   "Carrier_14_SpareInput(4_14)" AT %I1067.4 : Bool;   // SPARE INPUT
   "Carrier_14_SpareInput(4_15)" AT %I1067.5 : Bool;   // SPARE INPUT
   "Carrier_14_SpareInput(4_16)" AT %I1067.6 : Bool;   // SPARE INPUT
   "Carrier_14_SpareInput(4_17)" AT %I1067.7 : Bool;   // SPARE INPUT
   "Carrier_14_Slot5_Output" AT %IW1068 : Word;   // SLOT 5 OUTPUT WORD
   "Carrier_14_IRD400_HMI_24VDC_ENABLE" AT %I1068.0 : Bool;   // IRD 400 PANEL HMI 24V DC POWER
   "Carrier_14_FaultLight_LH" AT %I1068.1 : Bool;   // FAULT LIGHT LH
   "Carrier_14_RunLight_LH" AT %I1068.2 : Bool;   // RUN LIGHT LH
   "Carrier_14_FaultLight_RH" AT %I1068.3 : Bool;   // FAULT LIGHT RH
   "Carrier_14_RunLight_RH" AT %I1068.4 : Bool;   // RUN LIGHT RH
   "Carrier_14_SpareOutput(5_5)" AT %I1068.5 : Bool;   // SPARE OUTPUT
   "Carrier_14_SpareOutput(5_6)" AT %I1068.6 : Bool;   // SPARE OUTPUT
   "Carrier_14_SpareOutput(5_7)" AT %I1068.7 : Bool;   // SPARE OUTPUT
   "Carrier_14_ActualSpeed" AT %IW1070 : Word;   // ACTUAL SPEED
   "Carrier_14_CarrierDriveAlarm" AT %IW1072 : Word;   // CARRIER DRIVE ALARM
   "Carrier_14_CarrierDriveWarning" AT %IW1074 : Word;   // CARRIER DRIVE WARNING
   "Carrier_15_Status" AT %IW1100 : Word;   // CARRIER STATUS WORD
   "Carrier_15_Status.0" AT %I1100.0 : Bool;   // HEARTBEAT
   "Carrier_15_Status.1" AT %I1100.1 : Bool;   // MANUAL
   "Carrier_15_Status.2" AT %I1100.2 : Bool;   // IN_AUTO
   "Carrier_15_Status.3" AT %I1100.3 : Bool;   // POSITIONING_COMPLETE
   "Carrier_15_Status.4" AT %I1100.4 : Bool;   // PRODUCTION HOLD
   "Carrier_15_Status.5" AT %I1100.5 : Bool;   // CARRIER MOVING FORWARD
   "Carrier_15_Status.6" AT %I1100.6 : Bool;   // CARRIER MOVING REVERSE
   "Carrier_15_Status.7" AT %I1100.7 : Bool;   // CARRIER FAULT
   "Carrier_15_Status.8" AT %I1101.0 : Bool;   // CRASH DETECT TRIPPED
   "Carrier_15_Status.9" AT %I1101.1 : Bool;
   "Carrier_15_Status.10" AT %I1101.2 : Bool;
   "Carrier_15_Status.11" AT %I1101.3 : Bool;
   "Carrier_15_Status.12" AT %I1101.4 : Bool;
   "Carrier_15_Status.13" AT %I1101.5 : Bool;
   "Carrier_15_Status.14" AT %I1101.6 : Bool;
   "Carrier_15_Status.15" AT %I1101.7 : Bool;
   "Carrier_15_SDCFaultCode" AT %IW1102 : Word;   // SDC FAULT CODE
   "Carrier_15_CarrierPosition" AT %ID1104 : DWord;   // CARRIER POSITION
   "Carrier_15_CarrierNumber" AT %IW1108 : Word;   // CARRIER NUMBER
   "Carrier_15_G120DControlWord" AT %IW1111 : Word;   // G120D_STW1_CONTROL
   "Carrier_15_G120DControlWord.0" AT %I1111.0 : Bool;   // Bit_00_ON
   "Carrier_15_G120DControlWord.1" AT %I1111.1 : Bool;   // Bit_01_AUS2_INH
   "Carrier_15_G120DControlWord.2" AT %I1111.2 : Bool;   // Bit_02_AUS3_STOP
   "Carrier_15_G120DControlWord.3" AT %I1111.3 : Bool;   // Bit_03_EN
   "Carrier_15_G120DControlWord.4" AT %I1111.4 : Bool;   // Bit_04_EN_RAMP
   "Carrier_15_G120DControlWord.5" AT %I1111.5 : Bool;   // Bit_05_START_RAMP
   "Carrier_15_G120DControlWord.6" AT %I1111.6 : Bool;   // Bit_06_SETPOINT
   "Carrier_15_G120DControlWord.7" AT %I1111.7 : Bool;   // Bit_07_RESET
   "Carrier_15_G120DControlWord.8" AT %I1111.0 : Bool;   // Bit_08_JOG_R
   "Carrier_15_G120DControlWord.9" AT %I1111.1 : Bool;   // Bit_09_JOG_L
   "Carrier_15_G120DControlWord.10" AT %I1111.2 : Bool;   // Bit_10_CONTR_PLC
   "Carrier_15_G120DControlWord.11" AT %I1111.3 : Bool;   // Bit_11_REVERSE
   "Carrier_15_G120DControlWord.12" AT %I1111.4 : Bool;   // Bit_12_BRAKE_RELEASE
   "Carrier_15_G120DControlWord.13" AT %I1111.5 : Bool;   // Bit_13_DDS
   "Carrier_15_G120DControlWord.14" AT %I1111.6 : Bool;   // Bit_14_DO0
   "Carrier_15_G120DControlWord.15" AT %I1111.7 : Bool;   // Bit_15_DO1
   "Carrier_15_G120DStatusWord" AT %IW1112 : Word;   // G120D_ZSW1_STATUS
   "Carrier_15_G120DStatusWord.0" AT %I1112.0 : Bool;   // Bit_00_READY_RUN
   "Carrier_15_G120DStatusWord.1" AT %I1112.1 : Bool;   // Bit_01_READY_ON
   "Carrier_15_G120DStatusWord.2" AT %I1112.2 : Bool;   // Bit_02_ENABLE
   "Carrier_15_G120DStatusWord.3" AT %I1112.3 : Bool;   // Bit_03_FAULT
   "Carrier_15_G120DStatusWord.4" AT %I1112.4 : Bool;   // Bit_04_OFF2
   "Carrier_15_G120DStatusWord.5" AT %I1112.5 : Bool;   // Bit_05_OFF3
   "Carrier_15_G120DStatusWord.6" AT %I1112.6 : Bool;   // Bit_06_LOCK_OUT
   "Carrier_15_G120DStatusWord.7" AT %I1112.7 : Bool;   // Bit_07_WARN
   "Carrier_15_G120DStatusWord.8" AT %I1113.0 : Bool;   // Bit_08_NO_DEVIATION
   "Carrier_15_G120DStatusWord.9" AT %I1113.1 : Bool;   // Bit_09_CONTR_PLC
   "Carrier_15_G120DStatusWord.10" AT %I1113.2 : Bool;   // Bit_10_F_MAX
   "Carrier_15_G120DStatusWord.11" AT %I1113.3 : Bool;   // Bit_11_LIMIT_REACHED
   "Carrier_15_G120DStatusWord.12" AT %I1113.4 : Bool;   // Bit_12_BRAKE_OPEN
   "Carrier_15_G120DStatusWord.13" AT %I1113.5 : Bool;   // Bit_13_NO_OVERTEMP
   "Carrier_15_G120DStatusWord.14" AT %I1113.6 : Bool;   // Bit_14_CW_CCW
   "Carrier_15_G120DStatusWord.15" AT %I1113.7 : Bool;   // Bit_15_OVERL
   "Carrier_15_Slot2_Input" AT %IW1114 : Word;   // SLOT 2 INPUT WORD
   "Carrier_15_CrashDetectSW" AT %I1114.0 : Bool;   // CRASH DETECT SW
   "Carrier_15_SpareSafetyInput(2_1)" AT %I1114.1 : Bool;   // SPARE SAFETY INPUT
   "Carrier_15_SpareSafetyInput(2_2)" AT %I1114.2 : Bool;   // SPARE SAFETY INPUT
   "Carrier_15_SpareSafetyInput(2_3)" AT %I1114.3 : Bool;   // SPARE SAFETY INPUT
   "Carrier_15_SpareSafetyInput(2_4)" AT %I1114.4 : Bool;   // SPARE SAFETY INPUT
   "Carrier_15_SpareSafetyInput(2_5)" AT %I1114.5 : Bool;   // SPARE SAFETY INPUT
   "Carrier_15_SpareSafetyInput(2_6)" AT %I1114.6 : Bool;   // SPARE SAFETY INPUT
   "Carrier_15_SpareSafetyInput(2_7)" AT %I1114.7 : Bool;   // SPARE SAFETY INPUT
   "Carrier_15_Slot3_SafetyOutput" AT %IW1115 : Word;   // SLOT 3 SAFETY OUTPUT WORD
   "Carrier_15_Crash_Detect_OK" AT %I1115.0 : Bool;   // CARRIER CRASH DETECT
   "Carrier_15_SpareSafetyOutput(3_1)" AT %I1115.1 : Bool;   // SPARE SAFETY OUTPUT
   "Carrier_15_SpareSafetyOutput(3_2)" AT %I1115.2 : Bool;   // SPARE SAFETY OUTPUT
   "Carrier_15_SpareSafetyOutput(3_3)" AT %I1115.3 : Bool;   // SPARE SAFETY OUTPUT
   "Carrier_15_SpareSafetyOutput(3_4)" AT %I1115.4 : Bool;   // SPARE SAFETY OUTPUT
   "Carrier_15_SpareSafetyOutput(3_5)" AT %I1115.5 : Bool;   // SPARE SAFETY OUTPUT
   "Carrier_15_SpareSafetyOutput(3_6)" AT %I1115.6 : Bool;   // SPARE SAFETY OUTPUT
   "Carrier_15_SpareSafetyOutput(3_7)" AT %I1115.7 : Bool;   // SPARE SAFETY OUTPUT
   "Carrier_15_Slot4_Input" AT %IW1116 : Word;   // SLOT 4 INPUT WORD
   "Carrier_15_480VPowerOn_MDCB1" AT %I1116.0 : Bool;   // 480 VAC POWER ON MDCB 1
   "Carrier_15_SpareInput(4_1)" AT %I1116.1 : Bool;   // SPARE INPUT
   "Carrier_15_SpareInput(4_2)" AT %I1116.2 : Bool;   // SPARE INPUT
   "Carrier_15_SitopSelectStatus" AT %I1116.3 : Bool;   // SITOP SELECT STATUS
   "Carrier_15_DCsupplyOnPSCB2" AT %I1116.4 : Bool;   // DC SUPPLY ON PSCB 2
   "Carrier_15_SpareInput(4_5)" AT %I1116.5 : Bool;   // SPARE INPUT
   "Carrier_15_SpareInput(4_6)" AT %I1116.6 : Bool;   // SPARE INPUT
   "Carrier_15_SpareInput(4_7)" AT %I1116.7 : Bool;   // SPARE INPUT
   "Carrier_15_PB1_ProdHoldLH" AT %I1117.0 : Bool;   // PB 1 PRODUCTION HOLD LH
   "Carrier_15_PB2_ResetLH" AT %I1117.1 : Bool;   // PB 2 RESET LH
   "Carrier_15_PB3_ProdHoldRH" AT %I1117.2 : Bool;   // PB 3 PRODUCTION HOLD RH
   "Carrier_15_PB4_ResetRH" AT %I1117.3 : Bool;   // PB 4 RESET RH
   "Carrier_15_SpareInput(4_14)" AT %I1117.4 : Bool;   // SPARE INPUT
   "Carrier_15_SpareInput(4_15)" AT %I1117.5 : Bool;   // SPARE INPUT
   "Carrier_15_SpareInput(4_16)" AT %I1117.6 : Bool;   // SPARE INPUT
   "Carrier_15_SpareInput(4_17)" AT %I1117.7 : Bool;   // SPARE INPUT
   "Carrier_15_Slot5_Output" AT %IW1118 : Word;   // SLOT 5 OUTPUT WORD
   "Carrier_15_IRD400_HMI_24VDC_ENABLE" AT %I1118.0 : Bool;   // IRD 400 PANEL HMI 24V DC POWER
   "Carrier_15_FaultLight_LH" AT %I1118.1 : Bool;   // FAULT LIGHT LH
   "Carrier_15_RunLight_LH" AT %I1118.2 : Bool;   // RUN LIGHT LH
   "Carrier_15_FaultLight_RH" AT %I1118.3 : Bool;   // FAULT LIGHT RH
   "Carrier_15_RunLight_RH" AT %I1118.4 : Bool;   // RUN LIGHT RH
   "Carrier_15_SpareOutput(5_5)" AT %I1118.5 : Bool;   // SPARE OUTPUT
   "Carrier_15_SpareOutput(5_6)" AT %I1118.6 : Bool;   // SPARE OUTPUT
   "Carrier_15_SpareOutput(5_7)" AT %I1118.7 : Bool;   // SPARE OUTPUT
   "Carrier_15_ActualSpeed" AT %IW1120 : Word;   // ACTUAL SPEED
   "Carrier_15_CarrierDriveAlarm" AT %IW1122 : Word;   // CARRIER DRIVE ALARM
   "Carrier_15_CarrierDriveWarning" AT %IW1124 : Word;   // CARRIER DRIVE WARNING
   "Carrier_16_Status" AT %IW1150 : Word;   // CARRIER STATUS WORD
   "Carrier_16_Status.0" AT %I1150.0 : Bool;   // HEARTBEAT
   "Carrier_16_Status.1" AT %I1150.1 : Bool;   // MANUAL
   "Carrier_16_Status.2" AT %I1150.2 : Bool;   // IN_AUTO
   "Carrier_16_Status.3" AT %I1150.3 : Bool;   // POSITIONING_COMPLETE
   "Carrier_16_Status.4" AT %I1150.4 : Bool;   // PRODUCTION HOLD
   "Carrier_16_Status.5" AT %I1150.5 : Bool;   // CARRIER MOVING FORWARD
   "Carrier_16_Status.6" AT %I1150.6 : Bool;   // CARRIER MOVING REVERSE
   "Carrier_16_Status.7" AT %I1150.7 : Bool;   // CARRIER FAULT
   "Carrier_16_Status.8" AT %I1151.0 : Bool;   // CRASH DETECT TRIPPED
   "Carrier_16_Status.9" AT %I1151.1 : Bool;
   "Carrier_16_Status.10" AT %I1151.2 : Bool;
   "Carrier_16_Status.11" AT %I1151.3 : Bool;
   "Carrier_16_Status.12" AT %I1151.4 : Bool;
   "Carrier_16_Status.13" AT %I1151.5 : Bool;
   "Carrier_16_Status.14" AT %I1151.6 : Bool;
   "Carrier_16_Status.15" AT %I1151.7 : Bool;
   "Carrier_16_SDCFaultCode" AT %IW1152 : Word;   // SDC FAULT CODE
   "Carrier_16_CarrierPosition" AT %ID1154 : DWord;   // CARRIER POSITION
   "Carrier_16_CarrierNumber" AT %IW1158 : Word;   // CARRIER NUMBER
   "Carrier_16_G120DControlWord" AT %IW1160 : Word;   // G120D_STW1_CONTROL
   "Carrier_16_G120DControlWord.0" AT %I1160.0 : Bool;   // Bit_00_ON
   "Carrier_16_G120DControlWord.1" AT %I1160.1 : Bool;   // Bit_01_AUS2_INH
   "Carrier_16_G120DControlWord.2" AT %I1160.2 : Bool;   // Bit_02_AUS3_STOP
   "Carrier_16_G120DControlWord.3" AT %I1160.3 : Bool;   // Bit_03_EN
   "Carrier_16_G120DControlWord.4" AT %I1160.4 : Bool;   // Bit_04_EN_RAMP
   "Carrier_16_G120DControlWord.5" AT %I1160.5 : Bool;   // Bit_05_START_RAMP
   "Carrier_16_G120DControlWord.6" AT %I1160.6 : Bool;   // Bit_06_SETPOINT
   "Carrier_16_G120DControlWord.7" AT %I1160.7 : Bool;   // Bit_07_RESET
   "Carrier_16_G120DControlWord.8" AT %I1161.0 : Bool;   // Bit_08_JOG_R
   "Carrier_16_G120DControlWord.9" AT %I1161.1 : Bool;   // Bit_09_JOG_L
   "Carrier_16_G120DControlWord.10" AT %I1161.2 : Bool;   // Bit_10_CONTR_PLC
   "Carrier_16_G120DControlWord.11" AT %I1161.3 : Bool;   // Bit_11_REVERSE
   "Carrier_16_G120DControlWord.12" AT %I1161.4 : Bool;   // Bit_12_BRAKE_RELEASE
   "Carrier_16_G120DControlWord.13" AT %I1161.5 : Bool;   // Bit_13_DDS
   "Carrier_16_G120DControlWord.14" AT %I1161.6 : Bool;   // Bit_14_DO0
   "Carrier_16_G120DControlWord.15" AT %I1161.7 : Bool;   // Bit_15_DO1
   "Carrier_16_G120DStatusWord" AT %IW1162 : Word;   // G120D_ZSW1_STATUS
   "Carrier_16_G120DStatusWord.0" AT %I1162.0 : Bool;   // Bit_00_READY_RUN
   "Carrier_16_G120DStatusWord.1" AT %I1162.1 : Bool;   // Bit_01_READY_ON
   "Carrier_16_G120DStatusWord.2" AT %I1162.2 : Bool;   // Bit_02_ENABLE
   "Carrier_16_G120DStatusWord.3" AT %I1162.3 : Bool;   // Bit_03_FAULT
   "Carrier_16_G120DStatusWord.4" AT %I1162.4 : Bool;   // Bit_04_OFF2
   "Carrier_16_G120DStatusWord.5" AT %I1162.5 : Bool;   // Bit_05_OFF3
   "Carrier_16_G120DStatusWord.6" AT %I1162.6 : Bool;   // Bit_06_LOCK_OUT
   "Carrier_16_G120DStatusWord.7" AT %I1162.7 : Bool;   // Bit_07_WARN
   "Carrier_16_G120DStatusWord.8" AT %I1163.0 : Bool;   // Bit_08_NO_DEVIATION
   "Carrier_16_G120DStatusWord.9" AT %I1163.1 : Bool;   // Bit_09_CONTR_PLC
   "Carrier_16_G120DStatusWord.10" AT %I1163.2 : Bool;   // Bit_10_F_MAX
   "Carrier_16_G120DStatusWord.11" AT %I1163.3 : Bool;   // Bit_11_LIMIT_REACHED
   "Carrier_16_G120DStatusWord.12" AT %I1163.4 : Bool;   // Bit_12_BRAKE_OPEN
   "Carrier_16_G120DStatusWord.13" AT %I1163.5 : Bool;   // Bit_13_NO_OVERTEMP
   "Carrier_16_G120DStatusWord.14" AT %I1163.6 : Bool;   // Bit_14_CW_CCW
   "Carrier_16_G120DStatusWord.15" AT %I1163.7 : Bool;   // Bit_15_OVERL
   "Carrier_16_Slot2_Input" AT %IW1164 : Word;   // SLOT 2 INPUT WORD
   "Carrier_16_CrashDetectSW" AT %I1164.0 : Bool;   // CRASH DETECT SW
   "Carrier_16_SpareSafetyInput(2_1)" AT %I1164.1 : Bool;   // SPARE SAFETY INPUT
   "Carrier_16_SpareSafetyInput(2_2)" AT %I1164.2 : Bool;   // SPARE SAFETY INPUT
   "Carrier_16_SpareSafetyInput(2_3)" AT %I1164.3 : Bool;   // SPARE SAFETY INPUT
   "Carrier_16_SpareSafetyInput(2_4)" AT %I1164.4 : Bool;   // SPARE SAFETY INPUT
   "Carrier_16_SpareSafetyInput(2_5)" AT %I1164.5 : Bool;   // SPARE SAFETY INPUT
   "Carrier_16_SpareSafetyInput(2_6)" AT %I1164.6 : Bool;   // SPARE SAFETY INPUT
   "Carrier_16_SpareSafetyInput(2_7)" AT %I1164.7 : Bool;   // SPARE SAFETY INPUT
   "Carrier_16_Slot3_SafetyOutput" AT %IW1165 : Word;   // SLOT 3 SAFETY OUTPUT WORD
   "Carrier_16_Crash_Detect_OK" AT %I1165.0 : Bool;   // CARRIER CRASH DETECT
   "Carrier_16_SpareSafetyOutput(3_1)" AT %I1165.1 : Bool;   // SPARE SAFETY OUTPUT
   "Carrier_16_SpareSafetyOutput(3_2)" AT %I1165.2 : Bool;   // SPARE SAFETY OUTPUT
   "Carrier_16_SpareSafetyOutput(3_3)" AT %I1165.3 : Bool;   // SPARE SAFETY OUTPUT
   "Carrier_16_SpareSafetyOutput(3_4)" AT %I1165.4 : Bool;   // SPARE SAFETY OUTPUT
   "Carrier_16_SpareSafetyOutput(3_5)" AT %I1165.5 : Bool;   // SPARE SAFETY OUTPUT
   "Carrier_16_SpareSafetyOutput(3_6)" AT %I1165.6 : Bool;   // SPARE SAFETY OUTPUT
   "Carrier_16_SpareSafetyOutput(3_7)" AT %I1165.7 : Bool;   // SPARE SAFETY OUTPUT
   "Carrier_16_Slot4_Input" AT %IW1166 : Word;   // SLOT 4 INPUT WORD
   "Carrier_16_480VPowerOn_MDCB1" AT %I1166.0 : Bool;   // 480 VAC POWER ON MDCB 1
   "Carrier_16_SpareInput(4_1)" AT %I1166.1 : Bool;   // SPARE INPUT
   "Carrier_16_SpareInput(4_2)" AT %I1166.2 : Bool;   // SPARE INPUT
   "Carrier_16_SitopSelectStatus" AT %I1166.3 : Bool;   // SITOP SELECT STATUS
   "Carrier_16_DCsupplyOnPSCB2" AT %I1166.4 : Bool;   // DC SUPPLY ON PSCB 2
   "Carrier_16_SpareInput(4_5)" AT %I1166.5 : Bool;   // SPARE INPUT
   "Carrier_16_SpareInput(4_6)" AT %I1166.6 : Bool;   // SPARE INPUT
   "Carrier_16_SpareInput(4_7)" AT %I1166.7 : Bool;   // SPARE INPUT
   "Carrier_16_PB1_ProdHoldLH" AT %I1167.0 : Bool;   // PB 1 PRODUCTION HOLD LH
   "Carrier_16_PB2_ResetLH" AT %I1167.1 : Bool;   // PB 2 RESET LH
   "Carrier_16_PB3_ProdHoldRH" AT %I1167.2 : Bool;   // PB 3 PRODUCTION HOLD RH
   "Carrier_16_PB4_ResetRH" AT %I1167.3 : Bool;   // PB 4 RESET RH
   "Carrier_16_SpareInput(4_14)" AT %I1167.4 : Bool;   // SPARE INPUT
   "Carrier_16_SpareInput(4_15)" AT %I1167.5 : Bool;   // SPARE INPUT
   "Carrier_16_SpareInput(4_16)" AT %I1167.6 : Bool;   // SPARE INPUT
   "Carrier_16_SpareInput(4_17)" AT %I1167.7 : Bool;   // SPARE INPUT
   "Carrier_16_Slot5_Output" AT %IW1168 : Word;   // SLOT 5 OUTPUT WORD
   "Carrier_16_IRD400_HMI_24VDC_ENABLE" AT %I1168.0 : Bool;   // IRD 400 PANEL HMI 24V DC POWER
   "Carrier_16_FaultLight_LH" AT %I1168.1 : Bool;   // FAULT LIGHT LH
   "Carrier_16_RunLight_LH" AT %I1168.2 : Bool;   // RUN LIGHT LH
   "Carrier_16_FaultLight_RH" AT %I1168.3 : Bool;   // FAULT LIGHT RH
   "Carrier_16_RunLight_RH" AT %I1168.4 : Bool;   // RUN LIGHT RH
   "Carrier_16_SpareOutput(5_5)" AT %I1168.5 : Bool;   // SPARE OUTPUT
   "Carrier_16_SpareOutput(5_6)" AT %I1168.6 : Bool;   // SPARE OUTPUT
   "Carrier_16_SpareOutput(5_7)" AT %I1168.7 : Bool;   // SPARE OUTPUT
   "Carrier_16_ActualSpeed" AT %IW1170 : Word;   // ACTUAL SPEED
   "Carrier_16_CarrierDriveAlarm" AT %IW1172 : Word;   // CARRIER DRIVE ALARM
   "Carrier_16_CarrierDriveWarning" AT %IW1174 : Word;   // CARRIER DRIVE WARNING
   "Carrier_17_Status" AT %IW1200 : Word;   // CARRIER STATUS WORD
   "Carrier_17_Status.0" AT %I1200.0 : Bool;   // HEARTBEAT
   "Carrier_17_Status.1" AT %I1200.1 : Bool;   // MANUAL
   "Carrier_17_Status.2" AT %I1200.2 : Bool;   // IN_AUTO
   "Carrier_17_Status.3" AT %I1200.3 : Bool;   // POSITIONING_COMPLETE
   "Carrier_17_Status.4" AT %I1200.4 : Bool;   // PRODUCTION HOLD
   "Carrier_17_Status.5" AT %I1200.5 : Bool;   // CARRIER MOVING FORWARD
   "Carrier_17_Status.6" AT %I1200.6 : Bool;   // CARRIER MOVING REVERSE
   "Carrier_17_Status.7" AT %I1200.7 : Bool;   // CARRIER FAULT
   "Carrier_17_Status.8" AT %I1201.0 : Bool;   // CRASH DETECT TRIPPED
   "Carrier_17_Status.9" AT %I1201.1 : Bool;
   "Carrier_17_Status.10" AT %I1201.2 : Bool;
   "Carrier_17_Status.11" AT %I1201.3 : Bool;
   "Carrier_17_Status.12" AT %I1201.4 : Bool;
   "Carrier_17_Status.13" AT %I1201.5 : Bool;
   "Carrier_17_Status.14" AT %I1201.6 : Bool;
   "Carrier_17_Status.15" AT %I1201.7 : Bool;
   "Carrier_17_SDCFaultCode" AT %IW1202 : Word;   // SDC FAULT CODE
   "Carrier_17_CarrierPosition" AT %ID1204 : DWord;   // CARRIER POSITION
   "Carrier_17_CarrierNumber" AT %IW1208 : Word;   // CARRIER NUMBER
   "Carrier_17_G120DControlWord" AT %IW1212 : Word;   // G120D_STW1_CONTROL
   "Carrier_17_G120DControlWord.0" AT %I1212.0 : Bool;   // Bit_00_ON
   "Carrier_17_G120DControlWord.1" AT %I1212.1 : Bool;   // Bit_01_AUS2_INH
   "Carrier_17_G120DControlWord.2" AT %I1212.2 : Bool;   // Bit_02_AUS3_STOP
   "Carrier_17_G120DControlWord.3" AT %I1212.3 : Bool;   // Bit_03_EN
   "Carrier_17_G120DControlWord.4" AT %I1212.4 : Bool;   // Bit_04_EN_RAMP
   "Carrier_17_G120DControlWord.5" AT %I1212.5 : Bool;   // Bit_05_START_RAMP
   "Carrier_17_G120DControlWord.6" AT %I1212.6 : Bool;   // Bit_06_SETPOINT
   "Carrier_17_G120DControlWord.7" AT %I1212.7 : Bool;   // Bit_07_RESET
   "Carrier_17_G120DControlWord.8" AT %I1212.0 : Bool;   // Bit_08_JOG_R
   "Carrier_17_G120DControlWord.9" AT %I1212.1 : Bool;   // Bit_09_JOG_L
   "Carrier_17_G120DControlWord.10" AT %I1212.2 : Bool;   // Bit_10_CONTR_PLC
   "Carrier_17_G120DControlWord.11" AT %I1212.3 : Bool;   // Bit_11_REVERSE
   "Carrier_17_G120DControlWord.12" AT %I1212.4 : Bool;   // Bit_12_BRAKE_RELEASE
   "Carrier_17_G120DControlWord.13" AT %I1212.5 : Bool;   // Bit_13_DDS
   "Carrier_17_G120DControlWord.14" AT %I1212.6 : Bool;   // Bit_14_DO0
   "Carrier_17_G120DControlWord.15" AT %I1212.7 : Bool;   // Bit_15_DO1
   "Carrier_17_G120DStatusWord" AT %IW1212 : Word;   // G120D_ZSW1_STATUS
   "Carrier_17_G120DStatusWord.0" AT %I1212.0 : Bool;   // Bit_00_READY_RUN
   "Carrier_17_G120DStatusWord.1" AT %I1212.1 : Bool;   // Bit_01_READY_ON
   "Carrier_17_G120DStatusWord.2" AT %I1212.2 : Bool;   // Bit_02_ENABLE
   "Carrier_17_G120DStatusWord.3" AT %I1212.3 : Bool;   // Bit_03_FAULT
   "Carrier_17_G120DStatusWord.4" AT %I1212.4 : Bool;   // Bit_04_OFF2
   "Carrier_17_G120DStatusWord.5" AT %I1212.5 : Bool;   // Bit_05_OFF3
   "Carrier_17_G120DStatusWord.6" AT %I1212.6 : Bool;   // Bit_06_LOCK_OUT
   "Carrier_17_G120DStatusWord.7" AT %I1212.7 : Bool;   // Bit_07_WARN
   "Carrier_17_G120DStatusWord.8" AT %I1213.0 : Bool;   // Bit_08_NO_DEVIATION
   "Carrier_17_G120DStatusWord.9" AT %I1213.1 : Bool;   // Bit_09_CONTR_PLC
   "Carrier_17_G120DStatusWord.10" AT %I1213.2 : Bool;   // Bit_10_F_MAX
   "Carrier_17_G120DStatusWord.11" AT %I1213.3 : Bool;   // Bit_11_LIMIT_REACHED
   "Carrier_17_G120DStatusWord.12" AT %I1213.4 : Bool;   // Bit_12_BRAKE_OPEN
   "Carrier_17_G120DStatusWord.13" AT %I1213.5 : Bool;   // Bit_13_NO_OVERTEMP
   "Carrier_17_G120DStatusWord.14" AT %I1213.6 : Bool;   // Bit_14_CW_CCW
   "Carrier_17_G120DStatusWord.15" AT %I1213.7 : Bool;   // Bit_15_OVERL
   "Carrier_17_Slot2_Input" AT %IW1214 : Word;   // SLOT 2 INPUT WORD
   "Carrier_17_CrashDetectSW" AT %I1214.0 : Bool;   // CRASH DETECT SW
   "Carrier_17_SpareSafetyInput(2_1)" AT %I1214.1 : Bool;   // SPARE SAFETY INPUT
   "Carrier_17_SpareSafetyInput(2_2)" AT %I1214.2 : Bool;   // SPARE SAFETY INPUT
   "Carrier_17_SpareSafetyInput(2_3)" AT %I1214.3 : Bool;   // SPARE SAFETY INPUT
   "Carrier_17_SpareSafetyInput(2_4)" AT %I1214.4 : Bool;   // SPARE SAFETY INPUT
   "Carrier_17_SpareSafetyInput(2_5)" AT %I1214.5 : Bool;   // SPARE SAFETY INPUT
   "Carrier_17_SpareSafetyInput(2_6)" AT %I1214.6 : Bool;   // SPARE SAFETY INPUT
   "Carrier_17_SpareSafetyInput(2_7)" AT %I1214.7 : Bool;   // SPARE SAFETY INPUT
   "Carrier_17_Slot3_SafetyOutput" AT %IW1215 : Word;   // SLOT 3 SAFETY OUTPUT WORD
   "Carrier_17_Crash_Detect_OK" AT %I1215.0 : Bool;   // CARRIER CRASH DETECT
   "Carrier_17_SpareSafetyOutput(3_1)" AT %I1215.1 : Bool;   // SPARE SAFETY OUTPUT
   "Carrier_17_SpareSafetyOutput(3_2)" AT %I1215.2 : Bool;   // SPARE SAFETY OUTPUT
   "Carrier_17_SpareSafetyOutput(3_3)" AT %I1215.3 : Bool;   // SPARE SAFETY OUTPUT
   "Carrier_17_SpareSafetyOutput(3_4)" AT %I1215.4 : Bool;   // SPARE SAFETY OUTPUT
   "Carrier_17_SpareSafetyOutput(3_5)" AT %I1215.5 : Bool;   // SPARE SAFETY OUTPUT
   "Carrier_17_SpareSafetyOutput(3_6)" AT %I1215.6 : Bool;   // SPARE SAFETY OUTPUT
   "Carrier_17_SpareSafetyOutput(3_7)" AT %I1215.7 : Bool;   // SPARE SAFETY OUTPUT
   "Carrier_17_Slot4_Input" AT %IW1216 : Word;   // SLOT 4 INPUT WORD
   "Carrier_17_480VPowerOn_MDCB1" AT %I1216.0 : Bool;   // 480 VAC POWER ON MDCB 1
   "Carrier_17_SpareInput(4_1)" AT %I1216.1 : Bool;   // SPARE INPUT
   "Carrier_17_SpareInput(4_2)" AT %I1216.2 : Bool;   // SPARE INPUT
   "Carrier_17_SitopSelectStatus" AT %I1216.3 : Bool;   // SITOP SELECT STATUS
   "Carrier_17_DCsupplyOnPSCB2" AT %I1216.4 : Bool;   // DC SUPPLY ON PSCB 2
   "Carrier_17_SpareInput(4_5)" AT %I1216.5 : Bool;   // SPARE INPUT
   "Carrier_17_SpareInput(4_6)" AT %I1216.6 : Bool;   // SPARE INPUT
   "Carrier_17_SpareInput(4_7)" AT %I1216.7 : Bool;   // SPARE INPUT
   "Carrier_17_PB1_ProdHoldLH" AT %I1217.0 : Bool;   // PB 1 PRODUCTION HOLD LH
   "Carrier_17_PB2_ResetLH" AT %I1217.1 : Bool;   // PB 2 RESET LH
   "Carrier_17_PB3_ProdHoldRH" AT %I1217.2 : Bool;   // PB 3 PRODUCTION HOLD RH
   "Carrier_17_PB4_ResetRH" AT %I1217.3 : Bool;   // PB 4 RESET RH
   "Carrier_17_SpareInput(4_14)" AT %I1217.4 : Bool;   // SPARE INPUT
   "Carrier_17_SpareInput(4_15)" AT %I1217.5 : Bool;   // SPARE INPUT
   "Carrier_17_SpareInput(4_16)" AT %I1217.6 : Bool;   // SPARE INPUT
   "Carrier_17_SpareInput(4_17)" AT %I1217.7 : Bool;   // SPARE INPUT
   "Carrier_17_Slot5_Output" AT %IW1218 : Word;   // SLOT 5 OUTPUT WORD
   "Carrier_17_IRD400_HMI_24VDC_ENABLE" AT %I1218.0 : Bool;   // IRD 400 PANEL HMI 24V DC POWER
   "Carrier_17_FaultLight_LH" AT %I1218.1 : Bool;   // FAULT LIGHT LH
   "Carrier_17_RunLight_LH" AT %I1218.2 : Bool;   // RUN LIGHT LH
   "Carrier_17_FaultLight_RH" AT %I1218.3 : Bool;   // FAULT LIGHT RH
   "Carrier_17_RunLight_RH" AT %I1218.4 : Bool;   // RUN LIGHT RH
   "Carrier_17_SpareOutput(5_5)" AT %I1218.5 : Bool;   // SPARE OUTPUT
   "Carrier_17_SpareOutput(5_6)" AT %I1218.6 : Bool;   // SPARE OUTPUT
   "Carrier_17_SpareOutput(5_7)" AT %I1218.7 : Bool;   // SPARE OUTPUT
   "Carrier_17_ActualSpeed" AT %IW1220 : Word;   // ACTUAL SPEED
   "Carrier_17_CarrierDriveAlarm" AT %IW1222 : Word;   // CARRIER DRIVE ALARM
   "Carrier_17_CarrierDriveWarning" AT %IW1224 : Word;   // CARRIER DRIVE WARNING
   "Carrier_18_Status" AT %IW1250 : Word;   // CARRIER STATUS WORD
   "Carrier_18_Status.0" AT %I1250.0 : Bool;   // HEARTBEAT
   "Carrier_18_Status.1" AT %I1250.1 : Bool;   // MANUAL
   "Carrier_18_Status.2" AT %I1250.2 : Bool;   // IN_AUTO
   "Carrier_18_Status.3" AT %I1250.3 : Bool;   // POSITIONING_COMPLETE
   "Carrier_18_Status.4" AT %I1250.4 : Bool;   // PRODUCTION HOLD
   "Carrier_18_Status.5" AT %I1250.5 : Bool;   // CARRIER MOVING FORWARD
   "Carrier_18_Status.6" AT %I1250.6 : Bool;   // CARRIER MOVING REVERSE
   "Carrier_18_Status.7" AT %I1250.7 : Bool;   // CARRIER FAULT
   "Carrier_18_Status.8" AT %I1251.0 : Bool;   // CRASH DETECT TRIPPED
   "Carrier_18_Status.9" AT %I1251.1 : Bool;
   "Carrier_18_Status.10" AT %I1251.2 : Bool;
   "Carrier_18_Status.11" AT %I1251.3 : Bool;
   "Carrier_18_Status.12" AT %I1251.4 : Bool;
   "Carrier_18_Status.13" AT %I1251.5 : Bool;
   "Carrier_18_Status.14" AT %I1251.6 : Bool;
   "Carrier_18_Status.15" AT %I1251.7 : Bool;
   "Carrier_18_SDCFaultCode" AT %IW1252 : Word;   // SDC FAULT CODE
   "Carrier_18_CarrierPosition" AT %ID1254 : DWord;   // CARRIER POSITION
   "Carrier_18_CarrierNumber" AT %IW1258 : Word;   // CARRIER NUMBER
   "Carrier_18_G120DControlWord" AT %IW1260 : Word;   // G120D_STW1_CONTROL
   "Carrier_18_G120DControlWord.0" AT %I1260.0 : Bool;   // Bit_00_ON
   "Carrier_18_G120DControlWord.1" AT %I1260.1 : Bool;   // Bit_01_AUS2_INH
   "Carrier_18_G120DControlWord.2" AT %I1260.2 : Bool;   // Bit_02_AUS3_STOP
   "Carrier_18_G120DControlWord.3" AT %I1260.3 : Bool;   // Bit_03_EN
   "Carrier_18_G120DControlWord.4" AT %I1260.4 : Bool;   // Bit_04_EN_RAMP
   "Carrier_18_G120DControlWord.5" AT %I1260.5 : Bool;   // Bit_05_START_RAMP
   "Carrier_18_G120DControlWord.6" AT %I1260.6 : Bool;   // Bit_06_SETPOINT
   "Carrier_18_G120DControlWord.7" AT %I1260.7 : Bool;   // Bit_07_RESET
   "Carrier_18_G120DControlWord.8" AT %I1261.0 : Bool;   // Bit_08_JOG_R
   "Carrier_18_G120DControlWord.9" AT %I1261.1 : Bool;   // Bit_09_JOG_L
   "Carrier_18_G120DControlWord.10" AT %I1261.2 : Bool;   // Bit_10_CONTR_PLC
   "Carrier_18_G120DControlWord.11" AT %I1261.3 : Bool;   // Bit_11_REVERSE
   "Carrier_18_G120DControlWord.12" AT %I1261.4 : Bool;   // Bit_12_BRAKE_RELEASE
   "Carrier_18_G120DControlWord.13" AT %I1261.5 : Bool;   // Bit_13_DDS
   "Carrier_18_G120DControlWord.14" AT %I1261.6 : Bool;   // Bit_14_DO0
   "Carrier_18_G120DControlWord.15" AT %I1261.7 : Bool;   // Bit_15_DO1
   "Carrier_18_G120DStatusWord" AT %IW1262 : Word;   // G120D_ZSW1_STATUS
   "Carrier_18_G120DStatusWord.0" AT %I1262.0 : Bool;   // Bit_00_READY_RUN
   "Carrier_18_G120DStatusWord.1" AT %I1262.1 : Bool;   // Bit_01_READY_ON
   "Carrier_18_G120DStatusWord.2" AT %I1262.2 : Bool;   // Bit_02_ENABLE
   "Carrier_18_G120DStatusWord.3" AT %I1262.3 : Bool;   // Bit_03_FAULT
   "Carrier_18_G120DStatusWord.4" AT %I1262.4 : Bool;   // Bit_04_OFF2
   "Carrier_18_G120DStatusWord.5" AT %I1262.5 : Bool;   // Bit_05_OFF3
   "Carrier_18_G120DStatusWord.6" AT %I1262.6 : Bool;   // Bit_06_LOCK_OUT
   "Carrier_18_G120DStatusWord.7" AT %I1262.7 : Bool;   // Bit_07_WARN
   "Carrier_18_G120DStatusWord.8" AT %I1263.0 : Bool;   // Bit_08_NO_DEVIATION
   "Carrier_18_G120DStatusWord.9" AT %I1263.1 : Bool;   // Bit_09_CONTR_PLC
   "Carrier_18_G120DStatusWord.10" AT %I1263.2 : Bool;   // Bit_10_F_MAX
   "Carrier_18_G120DStatusWord.11" AT %I1263.3 : Bool;   // Bit_11_LIMIT_REACHED
   "Carrier_18_G120DStatusWord.12" AT %I1263.4 : Bool;   // Bit_12_BRAKE_OPEN
   "Carrier_18_G120DStatusWord.13" AT %I1263.5 : Bool;   // Bit_13_NO_OVERTEMP
   "Carrier_18_G120DStatusWord.14" AT %I1263.6 : Bool;   // Bit_14_CW_CCW
   "Carrier_18_G120DStatusWord.15" AT %I1263.7 : Bool;   // Bit_15_OVERL
   "Carrier_18_Slot2_Input" AT %IW1264 : Word;   // SLOT 2 INPUT WORD
   "Carrier_18_CrashDetectSW" AT %I1264.0 : Bool;   // CRASH DETECT SW
   "Carrier_18_SpareSafetyInput(2_1)" AT %I1264.1 : Bool;   // SPARE SAFETY INPUT
   "Carrier_18_SpareSafetyInput(2_2)" AT %I1264.2 : Bool;   // SPARE SAFETY INPUT
   "Carrier_18_SpareSafetyInput(2_3)" AT %I1264.3 : Bool;   // SPARE SAFETY INPUT
   "Carrier_18_SpareSafetyInput(2_4)" AT %I1264.4 : Bool;   // SPARE SAFETY INPUT
   "Carrier_18_SpareSafetyInput(2_5)" AT %I1264.5 : Bool;   // SPARE SAFETY INPUT
   "Carrier_18_SpareSafetyInput(2_6)" AT %I1264.6 : Bool;   // SPARE SAFETY INPUT
   "Carrier_18_SpareSafetyInput(2_7)" AT %I1264.7 : Bool;   // SPARE SAFETY INPUT
   "Carrier_18_Slot3_SafetyOutput" AT %IW1265 : Word;   // SLOT 3 SAFETY OUTPUT WORD
   "Carrier_18_Crash_Detect_OK" AT %I1265.0 : Bool;   // CARRIER CRASH DETECT
   "Carrier_18_SpareSafetyOutput(3_1)" AT %I1265.1 : Bool;   // SPARE SAFETY OUTPUT
   "Carrier_18_SpareSafetyOutput(3_2)" AT %I1265.2 : Bool;   // SPARE SAFETY OUTPUT
   "Carrier_18_SpareSafetyOutput(3_3)" AT %I1265.3 : Bool;   // SPARE SAFETY OUTPUT
   "Carrier_18_SpareSafetyOutput(3_4)" AT %I1265.4 : Bool;   // SPARE SAFETY OUTPUT
   "Carrier_18_SpareSafetyOutput(3_5)" AT %I1265.5 : Bool;   // SPARE SAFETY OUTPUT
   "Carrier_18_SpareSafetyOutput(3_6)" AT %I1265.6 : Bool;   // SPARE SAFETY OUTPUT
   "Carrier_18_SpareSafetyOutput(3_7)" AT %I1265.7 : Bool;   // SPARE SAFETY OUTPUT
   "Carrier_18_Slot4_Input" AT %IW1266 : Word;   // SLOT 4 INPUT WORD
   "Carrier_18_480VPowerOn_MDCB1" AT %I1266.0 : Bool;   // 480 VAC POWER ON MDCB 1
   "Carrier_18_SpareInput(4_1)" AT %I1266.1 : Bool;   // SPARE INPUT
   "Carrier_18_SpareInput(4_2)" AT %I1266.2 : Bool;   // SPARE INPUT
   "Carrier_18_SitopSelectStatus" AT %I1266.3 : Bool;   // SITOP SELECT STATUS
   "Carrier_18_DCsupplyOnPSCB2" AT %I1266.4 : Bool;   // DC SUPPLY ON PSCB 2
   "Carrier_18_SpareInput(4_5)" AT %I1266.5 : Bool;   // SPARE INPUT
   "Carrier_18_SpareInput(4_6)" AT %I1266.6 : Bool;   // SPARE INPUT
   "Carrier_18_SpareInput(4_7)" AT %I1266.7 : Bool;   // SPARE INPUT
   "Carrier_18_PB1_ProdHoldLH" AT %I1267.0 : Bool;   // PB 1 PRODUCTION HOLD LH
   "Carrier_18_PB2_ResetLH" AT %I1267.1 : Bool;   // PB 2 RESET LH
   "Carrier_18_PB3_ProdHoldRH" AT %I1267.2 : Bool;   // PB 3 PRODUCTION HOLD RH
   "Carrier_18_PB4_ResetRH" AT %I1267.3 : Bool;   // PB 4 RESET RH
   "Carrier_18_SpareInput(4_14)" AT %I1267.4 : Bool;   // SPARE INPUT
   "Carrier_18_SpareInput(4_15)" AT %I1267.5 : Bool;   // SPARE INPUT
   "Carrier_18_SpareInput(4_16)" AT %I1267.6 : Bool;   // SPARE INPUT
   "Carrier_18_SpareInput(4_17)" AT %I1267.7 : Bool;   // SPARE INPUT
   "Carrier_18_Slot5_Output" AT %IW1268 : Word;   // SLOT 5 OUTPUT WORD
   "Carrier_18_IRD400_HMI_24VDC_ENABLE" AT %I1268.0 : Bool;   // IRD 400 PANEL HMI 24V DC POWER
   "Carrier_18_FaultLight_LH" AT %I1268.1 : Bool;   // FAULT LIGHT LH
   "Carrier_18_RunLight_LH" AT %I1268.2 : Bool;   // RUN LIGHT LH
   "Carrier_18_FaultLight_RH" AT %I1268.3 : Bool;   // FAULT LIGHT RH
   "Carrier_18_RunLight_RH" AT %I1268.4 : Bool;   // RUN LIGHT RH
   "Carrier_18_SpareOutput(5_5)" AT %I1268.5 : Bool;   // SPARE OUTPUT
   "Carrier_18_SpareOutput(5_6)" AT %I1268.6 : Bool;   // SPARE OUTPUT
   "Carrier_18_SpareOutput(5_7)" AT %I1268.7 : Bool;   // SPARE OUTPUT
   "Carrier_18_ActualSpeed" AT %IW1270 : Word;   // ACTUAL SPEED
   "Carrier_18_CarrierDriveAlarm" AT %IW1272 : Word;   // CARRIER DRIVE ALARM
   "Carrier_18_CarrierDriveWarning" AT %IW1274 : Word;   // CARRIER DRIVE WARNING
   "Carrier_19_Status" AT %IW1300 : Word;   // CARRIER STATUS WORD
   "Carrier_19_Status.0" AT %I1300.0 : Bool;   // HEARTBEAT
   "Carrier_19_Status.1" AT %I1300.1 : Bool;   // MANUAL
   "Carrier_19_Status.2" AT %I1300.2 : Bool;   // IN_AUTO
   "Carrier_19_Status.3" AT %I1300.3 : Bool;   // POSITIONING_COMPLETE
   "Carrier_19_Status.4" AT %I1300.4 : Bool;   // PRODUCTION HOLD
   "Carrier_19_Status.5" AT %I1300.5 : Bool;   // CARRIER MOVING FORWARD
   "Carrier_19_Status.6" AT %I1300.6 : Bool;   // CARRIER MOVING REVERSE
   "Carrier_19_Status.7" AT %I1300.7 : Bool;   // CARRIER FAULT
   "Carrier_19_Status.8" AT %I1301.0 : Bool;   // CRASH DETECT TRIPPED
   "Carrier_19_Status.9" AT %I1301.1 : Bool;
   "Carrier_19_Status.10" AT %I1301.2 : Bool;
   "Carrier_19_Status.11" AT %I1301.3 : Bool;
   "Carrier_19_Status.12" AT %I1301.4 : Bool;
   "Carrier_19_Status.13" AT %I1301.5 : Bool;
   "Carrier_19_Status.14" AT %I1301.6 : Bool;
   "Carrier_19_Status.15" AT %I1301.7 : Bool;
   "Carrier_19_SDCFaultCode" AT %IW1302 : Word;   // SDC FAULT CODE
   "Carrier_19_CarrierPosition" AT %ID1304 : DWord;   // CARRIER POSITION
   "Carrier_19_CarrierNumber" AT %IW1308 : Word;   // CARRIER NUMBER
   "Carrier_19_G120DControlWord" AT %IW1310 : Word;   // G120D_STW1_CONTROL
   "Carrier_19_G120DControlWord.0" AT %I1310.0 : Bool;   // Bit_00_ON
   "Carrier_19_G120DControlWord.1" AT %I1310.1 : Bool;   // Bit_01_AUS2_INH
   "Carrier_19_G120DControlWord.2" AT %I1310.2 : Bool;   // Bit_02_AUS3_STOP
   "Carrier_19_G120DControlWord.3" AT %I1310.3 : Bool;   // Bit_03_EN
   "Carrier_19_G120DControlWord.4" AT %I1310.4 : Bool;   // Bit_04_EN_RAMP
   "Carrier_19_G120DControlWord.5" AT %I1310.5 : Bool;   // Bit_05_START_RAMP
   "Carrier_19_G120DControlWord.6" AT %I1310.6 : Bool;   // Bit_06_SETPOINT
   "Carrier_19_G120DControlWord.7" AT %I1310.7 : Bool;   // Bit_07_RESET
   "Carrier_19_G120DControlWord.8" AT %I1311.0 : Bool;   // Bit_08_JOG_R
   "Carrier_19_G120DControlWord.9" AT %I1311.1 : Bool;   // Bit_09_JOG_L
   "Carrier_19_G120DControlWord.10" AT %I1311.2 : Bool;   // Bit_10_CONTR_PLC
   "Carrier_19_G120DControlWord.11" AT %I1311.3 : Bool;   // Bit_11_REVERSE
   "Carrier_19_G120DControlWord.12" AT %I1311.4 : Bool;   // Bit_12_BRAKE_RELEASE
   "Carrier_19_G120DControlWord.13" AT %I1311.5 : Bool;   // Bit_13_DDS
   "Carrier_19_G120DControlWord.14" AT %I1311.6 : Bool;   // Bit_14_DO0
   "Carrier_19_G120DControlWord.15" AT %I1311.7 : Bool;   // Bit_15_DO1
   "Carrier_19_G120DStatusWord" AT %IW1312 : Word;   // G120D_ZSW1_STATUS
   "Carrier_19_G120DStatusWord.0" AT %I1312.0 : Bool;   // Bit_00_READY_RUN
   "Carrier_19_G120DStatusWord.1" AT %I1312.1 : Bool;   // Bit_01_READY_ON
   "Carrier_19_G120DStatusWord.2" AT %I1312.2 : Bool;   // Bit_02_ENABLE
   "Carrier_19_G120DStatusWord.3" AT %I1312.3 : Bool;   // Bit_03_FAULT
   "Carrier_19_G120DStatusWord.4" AT %I1312.4 : Bool;   // Bit_04_OFF2
   "Carrier_19_G120DStatusWord.5" AT %I1312.5 : Bool;   // Bit_05_OFF3